   
   ////MSHIFTSBR
   	ELSIF (TMP_dSourceFile = 201) AND (TMP_dDestFile = 200) THEN
   		COP(N201[TMP_dSourceOffset], N200[TMP_dDestOffset], TMP_dNumValues);
   	ELSIF (TMP_dSourceFile = 202) AND (TMP_dDestFile = 200) THEN
   		COP(N202[TMP_dSourceOffset], N200[TMP_dDestOffset], TMP_dNumValues);
   	ELSIF (TMP_dSourceFile = 203) AND (TMP_dDestFile = 200) THEN
   		COP(N203[TMP_dSourceOffset], N200[TMP_dDestOffset], TMP_dNumValues);
   	ELSIF (TMP_dSourceFile = 204) AND (TMP_dDestFile = 200) THEN
   		COP(N204[TMP_dSourceOffset], N200[TMP_dDestOffset], TMP_dNumValues);
   	ELSIF (TMP_dSourceFile = 205) AND (TMP_dDestFile = 200) THEN
   		COP(N205[TMP_dSourceOffset], N200[TMP_dDestOffset], TMP_dNumValues);
   	ELSIF (TMP_dSourceFile = 206) AND (TMP_dDestFile = 200) THEN
   		COP(N206[TMP_dSourceOffset], N200[TMP_dDestOffset], TMP_dNumValues);
   	ELSIF (TMP_dSourceFile = 207) AND (TMP_dDestFile = 200) THEN
   		COP(N207[TMP_dSourceOffset], N200[TMP_dDestOffset], TMP_dNumValues);
   	ELSIF (TMP_dSourceFile = 208) AND (TMP_dDestFile = 200) THEN
   		COP(N208[TMP_dSourceOffset], N200[TMP_dDestOffset], TMP_dNumValues);
   	ELSIF (TMP_dSourceFile = 209) AND (TMP_dDestFile = 200) THEN
   		COP(N209[TMP_dSourceOffset], N200[TMP_dDestOffset], TMP_dNumValues);
   	ELSIF (TMP_dSourceFile = 210) AND (TMP_dDestFile = 200) THEN
   		COP(N210[TMP_dSourceOffset], N200[TMP_dDestOffset], TMP_dNumValues);
   	ELSIF (TMP_dSourceFile = 211) AND (TMP_dDestFile = 200) THEN
   		COP(N211[TMP_dSourceOffset], N200[TMP_dDestOffset], TMP_dNumValues);
   	ELSIF (TMP_dSourceFile = 212) AND (TMP_dDestFile = 200) THEN
   		COP(N212[TMP_dSourceOffset], N200[TMP_dDestOffset], TMP_dNumValues);
   	ELSIF (TMP_dSourceFile = 213) AND (TMP_dDestFile = 200) THEN
   		COP(N213[TMP_dSourceOffset], N200[TMP_dDestOffset], TMP_dNumValues);
   	ELSIF (TMP_dSourceFile = 214) AND (TMP_dDestFile = 200) THEN
   		COP(N214[TMP_dSourceOffset], N200[TMP_dDestOffset], TMP_dNumValues);
   	ELSIF (TMP_dSourceFile = 215) AND (TMP_dDestFile = 200) THEN
   		COP(N215[TMP_dSourceOffset], N200[TMP_dDestOffset], TMP_dNumValues);
   	ELSIF (TMP_dSourceFile = 216) AND (TMP_dDestFile = 200) THEN
   		COP(N216[TMP_dSourceOffset], N200[TMP_dDestOffset], TMP_dNumValues);
   	ELSIF (TMP_dSourceFile = 217) AND (TMP_dDestFile = 200) THEN
   		COP(N217[TMP_dSourceOffset], N200[TMP_dDestOffset], TMP_dNumValues);
   	ELSIF (TMP_dSourceFile = 218) AND (TMP_dDestFile = 200) THEN
   		COP(N218[TMP_dSourceOffset], N200[TMP_dDestOffset], TMP_dNumValues);
   
   	ELSIF (TMP_dSourceFile = 200) AND (TMP_dDestFile = 201) THEN
   		COP(N200[TMP_dSourceOffset], N201[TMP_dDestOffset], TMP_dNumValues);
   	ELSIF (TMP_dSourceFile = 200) AND (TMP_dDestFile = 202) THEN
   		COP(N200[TMP_dSourceOffset], N202[TMP_dDestOffset], TMP_dNumValues);
   	ELSIF (TMP_dSourceFile = 200) AND (TMP_dDestFile = 203) THEN
   		COP(N200[TMP_dSourceOffset], N203[TMP_dDestOffset], TMP_dNumValues);
   	ELSIF (TMP_dSourceFile = 200) AND (TMP_dDestFile = 204) THEN
   		COP(N200[TMP_dSourceOffset], N204[TMP_dDestOffset], TMP_dNumValues);
   	ELSIF (TMP_dSourceFile = 200) AND (TMP_dDestFile = 205) THEN
   		COP(N200[TMP_dSourceOffset], N205[TMP_dDestOffset], TMP_dNumValues);
   	ELSIF (TMP_dSourceFile = 200) AND (TMP_dDestFile = 206) THEN
   		COP(N200[TMP_dSourceOffset], N206[TMP_dDestOffset], TMP_dNumValues);
   	ELSIF (TMP_dSourceFile = 200) AND (TMP_dDestFile = 207) THEN
   		COP(N200[TMP_dSourceOffset], N207[TMP_dDestOffset], TMP_dNumValues);
   	ELSIF (TMP_dSourceFile = 200) AND (TMP_dDestFile = 208) THEN
   		COP(N200[TMP_dSourceOffset], N208[TMP_dDestOffset], TMP_dNumValues);
   	ELSIF (TMP_dSourceFile = 200) AND (TMP_dDestFile = 209) THEN
   		COP(N200[TMP_dSourceOffset], N209[TMP_dDestOffset], TMP_dNumValues);
   	ELSIF (TMP_dSourceFile = 200) AND (TMP_dDestFile = 210) THEN
   		COP(N200[TMP_dSourceOffset], N210[TMP_dDestOffset], TMP_dNumValues);
   	ELSIF (TMP_dSourceFile = 200) AND (TMP_dDestFile = 211) THEN
   		COP(N200[TMP_dSourceOffset], N211[TMP_dDestOffset], TMP_dNumValues);
   	ELSIF (TMP_dSourceFile = 200) AND (TMP_dDestFile = 212) THEN
   		COP(N200[TMP_dSourceOffset], N212[TMP_dDestOffset], TMP_dNumValues);
   	ELSIF (TMP_dSourceFile = 200) AND (TMP_dDestFile = 213) THEN
   		COP(N200[TMP_dSourceOffset], N213[TMP_dDestOffset], TMP_dNumValues);
   	ELSIF (TMP_dSourceFile = 200) AND (TMP_dDestFile = 214) THEN
   		COP(N200[TMP_dSourceOffset], N214[TMP_dDestOffset], TMP_dNumValues);
   	ELSIF (TMP_dSourceFile = 200) AND (TMP_dDestFile = 215) THEN
   		COP(N200[TMP_dSourceOffset], N215[TMP_dDestOffset], TMP_dNumValues);
   	ELSIF (TMP_dSourceFile = 200) AND (TMP_dDestFile = 216) THEN
   		COP(N200[TMP_dSourceOffset], N216[TMP_dDestOffset], TMP_dNumValues);
   	ELSIF (TMP_dSourceFile = 200) AND (TMP_dDestFile = 217) THEN
   		COP(N200[TMP_dSourceOffset], N217[TMP_dDestOffset], TMP_dNumValues);
   	ELSIF (TMP_dSourceFile = 200) AND (TMP_dDestFile = 218) THEN
   		COP(N200[TMP_dSourceOffset], N218[TMP_dDestOffset], TMP_dNumValues);
   
   
   ////////
   	ELSE
   		TMP_dErrSourceFile := TMP_dSourceFile;
   		TMP_dErrDestFile := TMP_dDestFile;
   	END_IF;
   *)
   
   RET(TMP_dErrSourceFile,TMP_dErrDestFile);
   
END_ROUTINE

ROUTINE _9_MCP_H   (* ladder *)
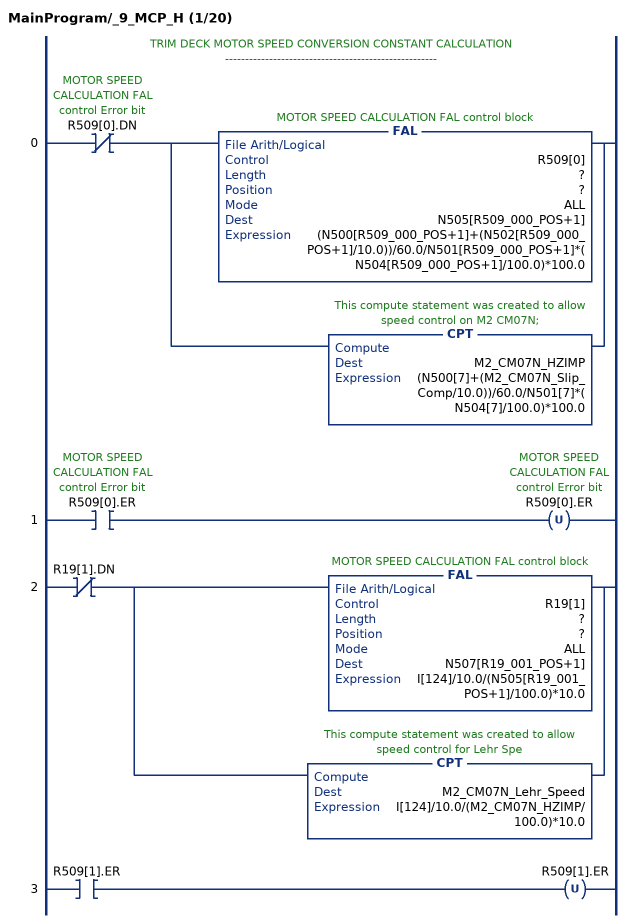
   // TRIM DECK MOTOR SPEED CONVERSION CONSTANT CALCULATION
   // -----------------------------------------------------
   0: XIO(R509[0].DN)[FAL(R509[0],?,?,ALL,N505[R509_000_POS+1],(N500[R509_000_POS+1]+(N502[R509_000_POS+1]/10.0))/60.0/N501[R509_000_POS+1]*(N504[R509_000_POS+1]/100.0)*100.0) ,CPT(M2_CM07N_HZIMP,(N500[7]+(M2_CM07N_Slip_Comp/10.0))/60.0/N501[7]*(N504[7]/100.0)*100.0) ];
   1: XIC(R509[0].ER)OTU(R509[0].ER);
   2: XIO(R19[1].DN)[FAL(R19[1],?,?,ALL,N507[R19_001_POS+1],I[124]/10.0/(N505[R19_001_POS+1]/100.0)*10.0) ,CPT(M2_CM07N_Lehr_Speed,I[124]/10.0/(M2_CM07N_HZIMP/100.0)*10.0) ];
   3: XIC(R509[1].ER)OTU(R509[1].ER);
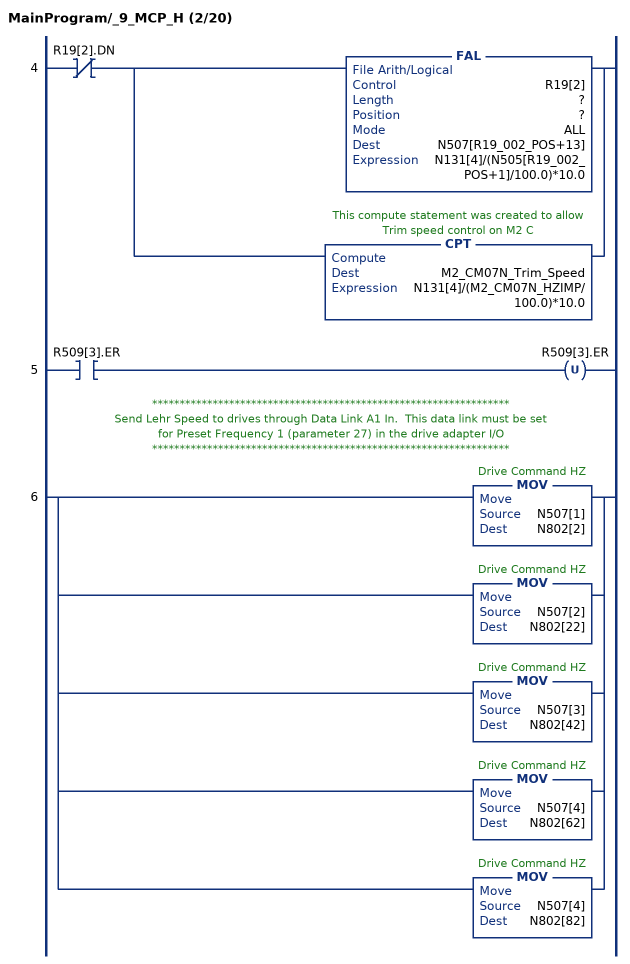
   4: XIO(R19[2].DN)[FAL(R19[2],?,?,ALL,N507[R19_002_POS+13],N131[4]/(N505[R19_002_POS+1]/100.0)*10.0) ,CPT(M2_CM07N_Trim_Speed,N131[4]/(M2_CM07N_HZIMP/100.0)*10.0) ];
   5: XIC(R509[3].ER)OTU(R509[3].ER);
   // *****************************************************************
   // Send Lehr Speed to drives through Data Link A1 In.  This data link must be set
   // for Preset Frequency 1 (parameter 27) in the drive adapter I/O
   // *****************************************************************
   6: [MOV(N507[1],N802[2]) ,MOV(N507[2],N802[22]) ,MOV(N507[3],N802[42]) ,MOV(N507[4],N802[62]) ,MOV(N507[4],N802[82]) ];
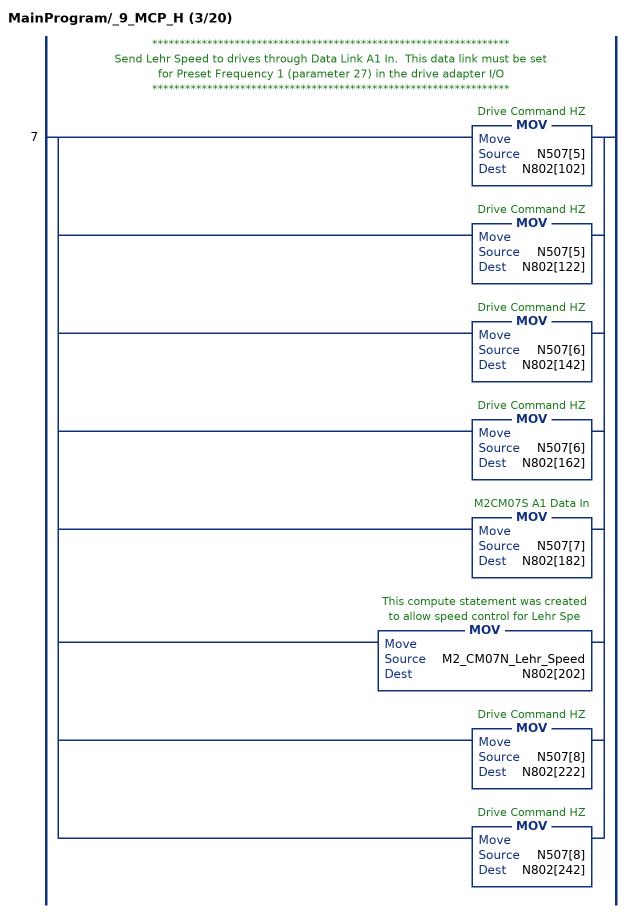
   // *****************************************************************
   // Send Lehr Speed to drives through Data Link A1 In.  This data link must be set
   // for Preset Frequency 1 (parameter 27) in the drive adapter I/O
   // *****************************************************************
   7: [MOV(N507[5],N802[102]) ,MOV(N507[5],N802[122]) ,MOV(N507[6],N802[142]) ,MOV(N507[6],N802[162]) ,MOV(N507[7],N802[182]) ,MOV(M2_CM07N_Lehr_Speed,N802[202]) ,MOV(N507[8],N802[222]) ,MOV(N507[8],N802[242]) ];
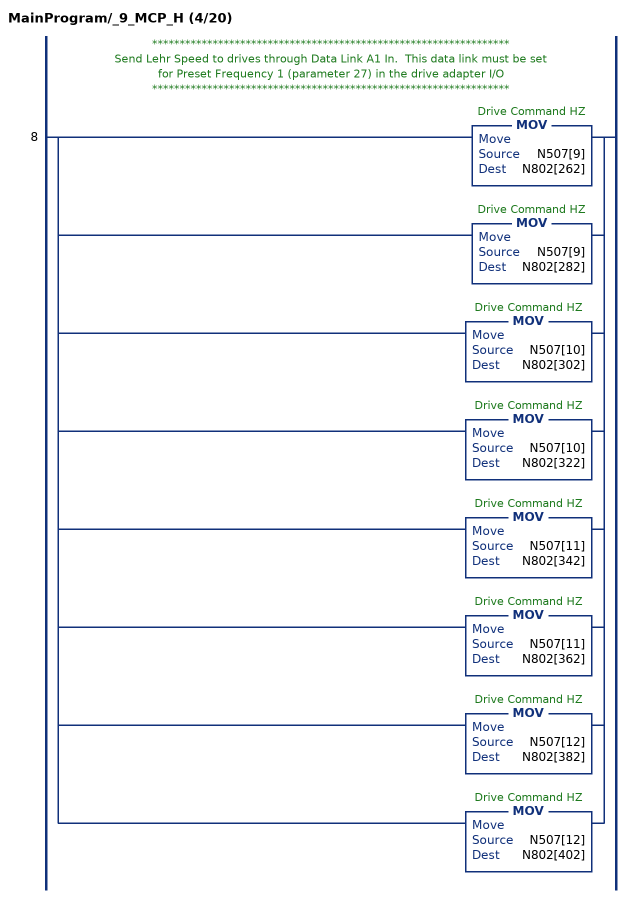
   // *****************************************************************
   // Send Lehr Speed to drives through Data Link A1 In.  This data link must be set
   // for Preset Frequency 1 (parameter 27) in the drive adapter I/O
   // *****************************************************************
   8: [MOV(N507[9],N802[262]) ,MOV(N507[9],N802[282]) ,MOV(N507[10],N802[302]) ,MOV(N507[10],N802[322]) ,MOV(N507[11],N802[342]) ,MOV(N507[11],N802[362]) ,MOV(N507[12],N802[382]) ,MOV(N507[12],N802[402]) ];
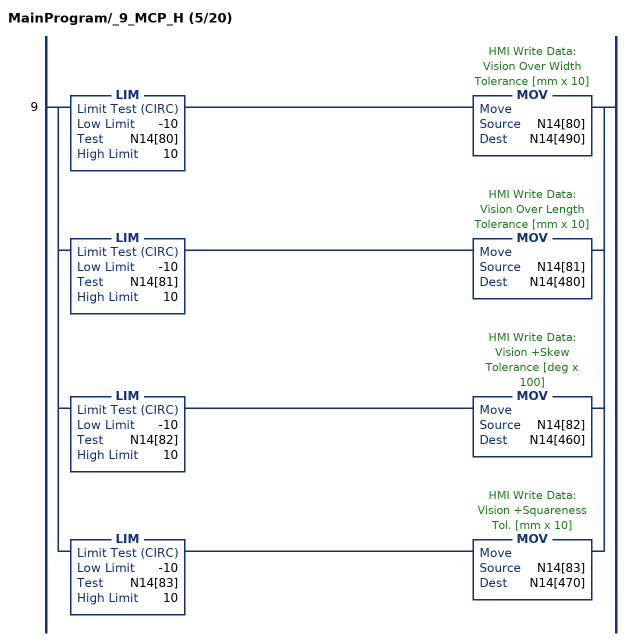
   9: [LIM(-10,N14[80],10) MOV(N14[80],N14[490]) ,LIM(-10,N14[81],10) MOV(N14[81],N14[480]) ,LIM(-10,N14[82],10) MOV(N14[82],N14[460]) ,LIM(-10,N14[83],10) MOV(N14[83],N14[470]) ];
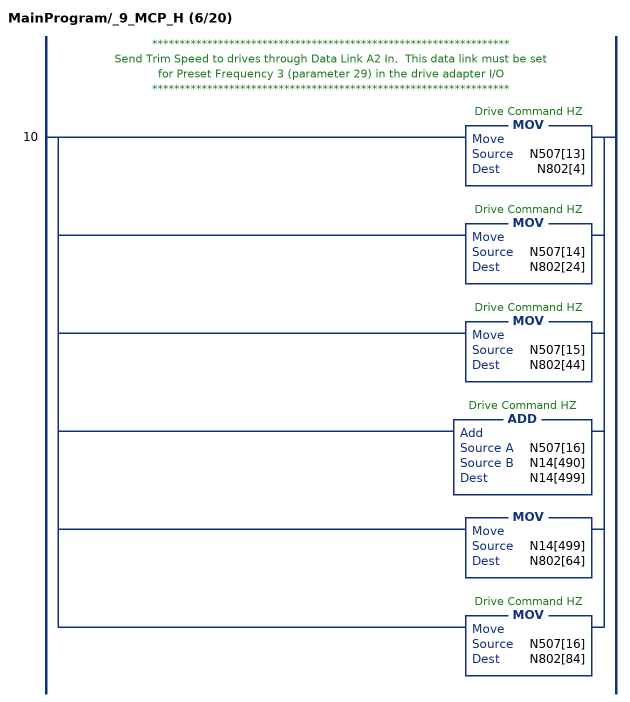
   // *****************************************************************
   // Send Trim Speed to drives through Data Link A2 In.  This data link must be set
   // for Preset Frequency 3 (parameter 29) in the drive adapter I/O
   // *****************************************************************
   10: [MOV(N507[13],N802[4]) ,MOV(N507[14],N802[24]) ,MOV(N507[15],N802[44]) ,ADD(N507[16],N14[490],N14[499]) ,MOV(N14[499],N802[64]) ,MOV(N507[16],N802[84]) ];
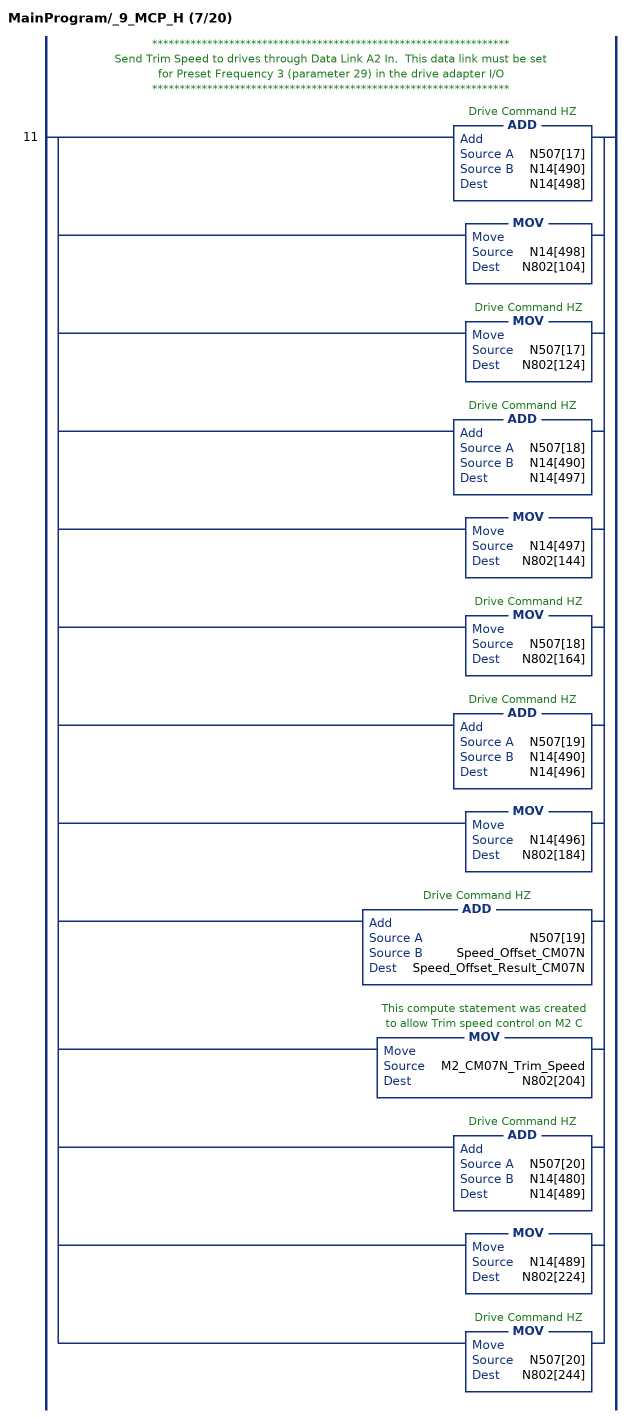
   // *****************************************************************
   // Send Trim Speed to drives through Data Link A2 In.  This data link must be set
   // for Preset Frequency 3 (parameter 29) in the drive adapter I/O
   // *****************************************************************
   11: [ADD(N507[17],N14[490],N14[498]) ,MOV(N14[498],N802[104]) ,MOV(N507[17],N802[124]) ,ADD(N507[18],N14[490],N14[497]) ,MOV(N14[497],N802[144]) ,MOV(N507[18],N802[164]) ,ADD(N507[19],N14[490],N14[496]) ,MOV(N14[496],N802[184]) ,ADD(N507[19],Speed_Offset_CM07N,Speed_Offset_Result_CM07N) ,MOV(M2_CM07N_Trim_Speed,N802[204]) ,ADD(N507[20],N14[480],N14[489]) ,MOV(N14[489],N802[224]) ,MOV(N507[20],N802[244]) ];
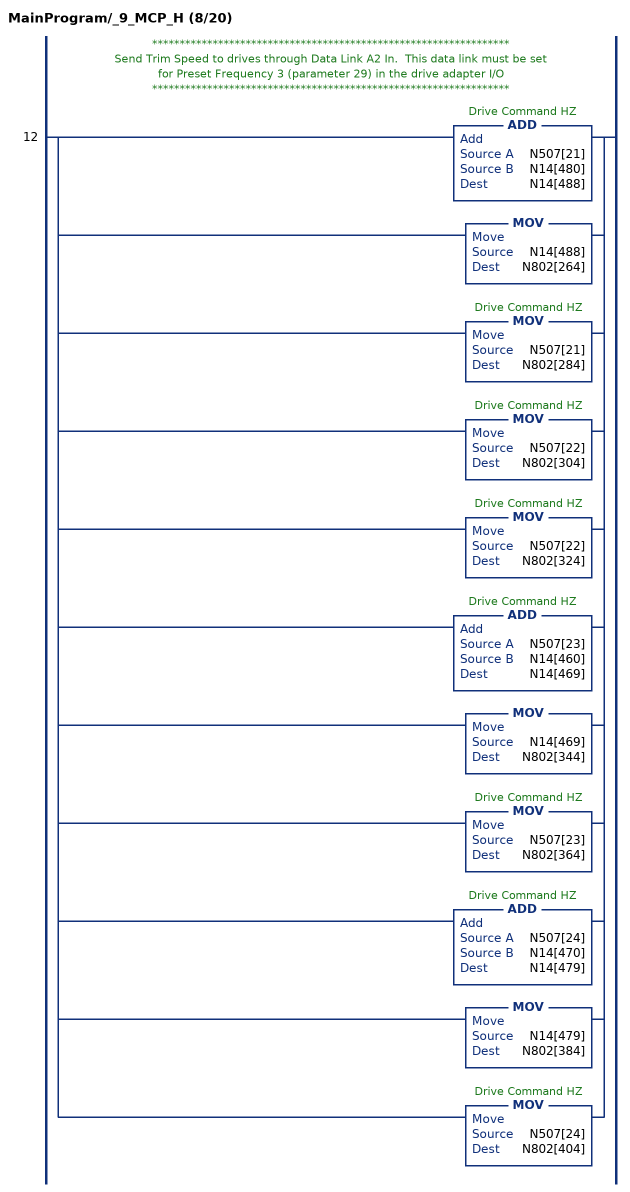
   // *****************************************************************
   // Send Trim Speed to drives through Data Link A2 In.  This data link must be set
   // for Preset Frequency 3 (parameter 29) in the drive adapter I/O
   // *****************************************************************
   12: [ADD(N507[21],N14[480],N14[488]) ,MOV(N14[488],N802[264]) ,MOV(N507[21],N802[284]) ,MOV(N507[22],N802[304]) ,MOV(N507[22],N802[324]) ,ADD(N507[23],N14[460],N14[469]) ,MOV(N14[469],N802[344]) ,MOV(N507[23],N802[364]) ,ADD(N507[24],N14[470],N14[479]) ,MOV(N14[479],N802[384]) ,MOV(N507[24],N802[404]) ];
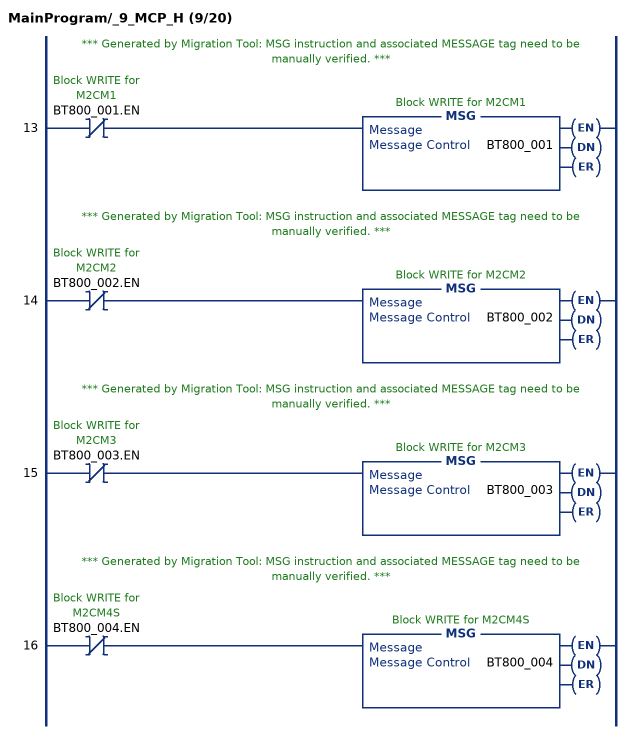
   // *** Generated by Migration Tool: MSG instruction and associated MESSAGE tag need to be manually verified. ***
   13: XIO(BT800_001.EN)MSG(BT800_001);
   // *** Generated by Migration Tool: MSG instruction and associated MESSAGE tag need to be manually verified. ***
   14: XIO(BT800_002.EN)MSG(BT800_002);
   // *** Generated by Migration Tool: MSG instruction and associated MESSAGE tag need to be manually verified. ***
   15: XIO(BT800_003.EN)MSG(BT800_003);
   // *** Generated by Migration Tool: MSG instruction and associated MESSAGE tag need to be manually verified. ***
   16: XIO(BT800_004.EN)MSG(BT800_004);
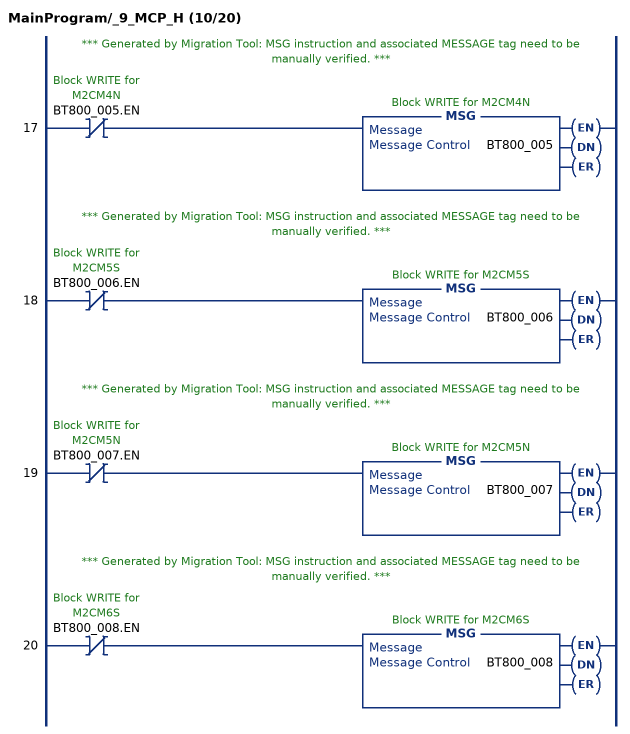
   // *** Generated by Migration Tool: MSG instruction and associated MESSAGE tag need to be manually verified. ***
   17: XIO(BT800_005.EN)MSG(BT800_005);
   // *** Generated by Migration Tool: MSG instruction and associated MESSAGE tag need to be manually verified. ***
   18: XIO(BT800_006.EN)MSG(BT800_006);
   // *** Generated by Migration Tool: MSG instruction and associated MESSAGE tag need to be manually verified. ***
   19: XIO(BT800_007.EN)MSG(BT800_007);
   // *** Generated by Migration Tool: MSG instruction and associated MESSAGE tag need to be manually verified. ***
   20: XIO(BT800_008.EN)MSG(BT800_008);
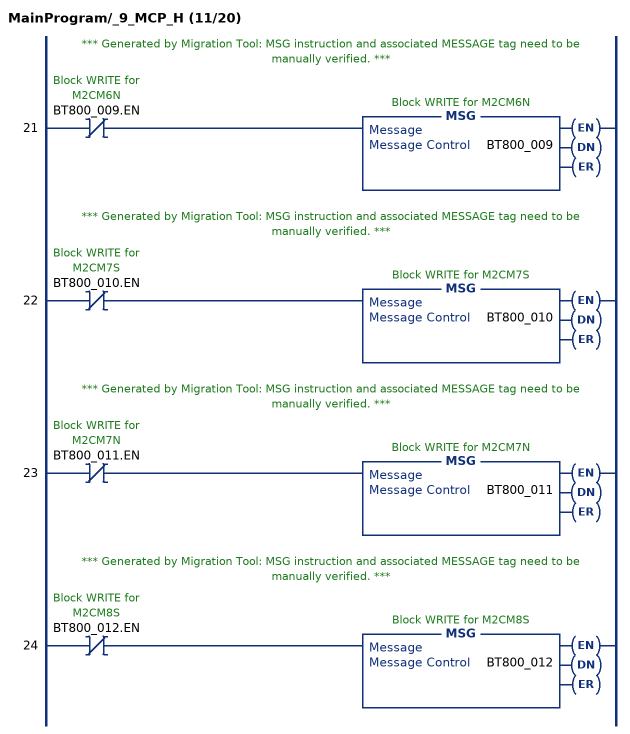
   // *** Generated by Migration Tool: MSG instruction and associated MESSAGE tag need to be manually verified. ***
   21: XIO(BT800_009.EN)MSG(BT800_009);
   // *** Generated by Migration Tool: MSG instruction and associated MESSAGE tag need to be manually verified. ***
   22: XIO(BT800_010.EN)MSG(BT800_010);
   // *** Generated by Migration Tool: MSG instruction and associated MESSAGE tag need to be manually verified. ***
   23: XIO(BT800_011.EN)MSG(BT800_011);
   // *** Generated by Migration Tool: MSG instruction and associated MESSAGE tag need to be manually verified. ***
   24: XIO(BT800_012.EN)MSG(BT800_012);
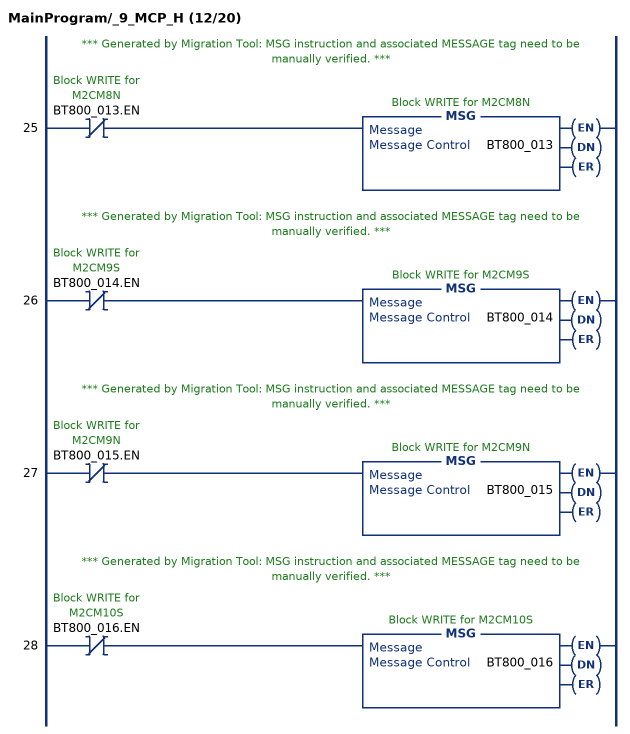
   // *** Generated by Migration Tool: MSG instruction and associated MESSAGE tag need to be manually verified. ***
   25: XIO(BT800_013.EN)MSG(BT800_013);
   // *** Generated by Migration Tool: MSG instruction and associated MESSAGE tag need to be manually verified. ***
   26: XIO(BT800_014.EN)MSG(BT800_014);
   // *** Generated by Migration Tool: MSG instruction and associated MESSAGE tag need to be manually verified. ***
   27: XIO(BT800_015.EN)MSG(BT800_015);
   // *** Generated by Migration Tool: MSG instruction and associated MESSAGE tag need to be manually verified. ***
   28: XIO(BT800_016.EN)MSG(BT800_016);
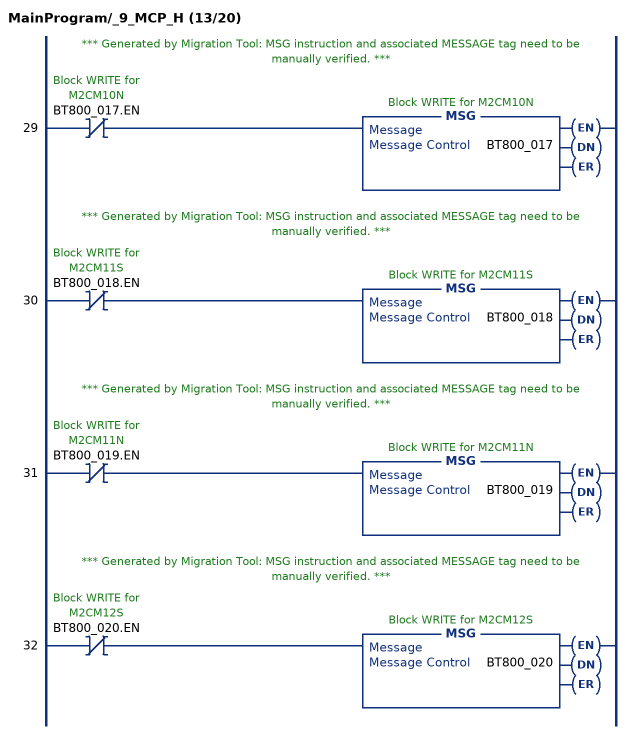
   // *** Generated by Migration Tool: MSG instruction and associated MESSAGE tag need to be manually verified. ***
   29: XIO(BT800_017.EN)MSG(BT800_017);
   // *** Generated by Migration Tool: MSG instruction and associated MESSAGE tag need to be manually verified. ***
   30: XIO(BT800_018.EN)MSG(BT800_018);
   // *** Generated by Migration Tool: MSG instruction and associated MESSAGE tag need to be manually verified. ***
   31: XIO(BT800_019.EN)MSG(BT800_019);
   // *** Generated by Migration Tool: MSG instruction and associated MESSAGE tag need to be manually verified. ***
   32: XIO(BT800_020.EN)MSG(BT800_020);
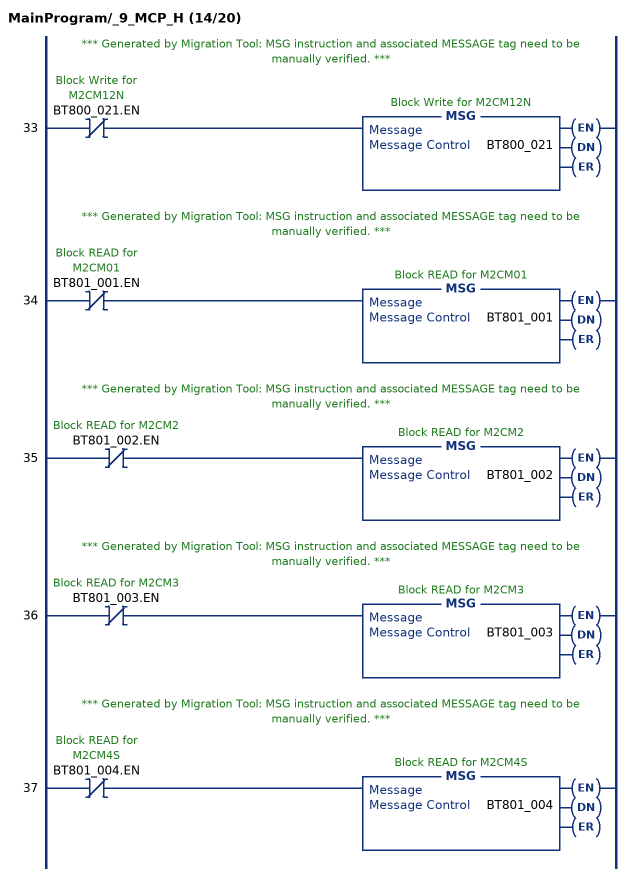
   // *** Generated by Migration Tool: MSG instruction and associated MESSAGE tag need to be manually verified. ***
   33: XIO(BT800_021.EN)MSG(BT800_021);
   // *** Generated by Migration Tool: MSG instruction and associated MESSAGE tag need to be manually verified. ***
   34: XIO(BT801_001.EN)MSG(BT801_001);
   // *** Generated by Migration Tool: MSG instruction and associated MESSAGE tag need to be manually verified. ***
   35: XIO(BT801_002.EN)MSG(BT801_002);
   // *** Generated by Migration Tool: MSG instruction and associated MESSAGE tag need to be manually verified. ***
   36: XIO(BT801_003.EN)MSG(BT801_003);
   // *** Generated by Migration Tool: MSG instruction and associated MESSAGE tag need to be manually verified. ***
   37: XIO(BT801_004.EN)MSG(BT801_004);
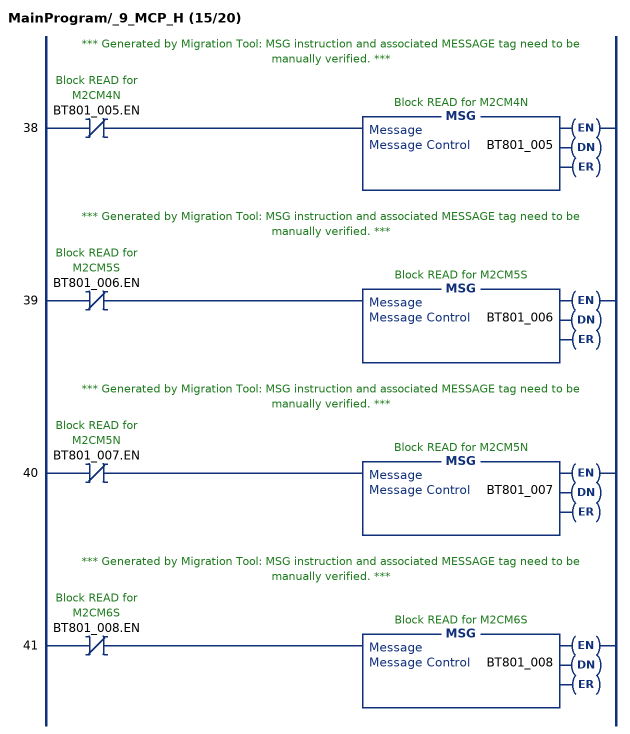
   // *** Generated by Migration Tool: MSG instruction and associated MESSAGE tag need to be manually verified. ***
   38: XIO(BT801_005.EN)MSG(BT801_005);
   // *** Generated by Migration Tool: MSG instruction and associated MESSAGE tag need to be manually verified. ***
   39: XIO(BT801_006.EN)MSG(BT801_006);
   // *** Generated by Migration Tool: MSG instruction and associated MESSAGE tag need to be manually verified. ***
   40: XIO(BT801_007.EN)MSG(BT801_007);
   // *** Generated by Migration Tool: MSG instruction and associated MESSAGE tag need to be manually verified. ***
   41: XIO(BT801_008.EN)MSG(BT801_008);
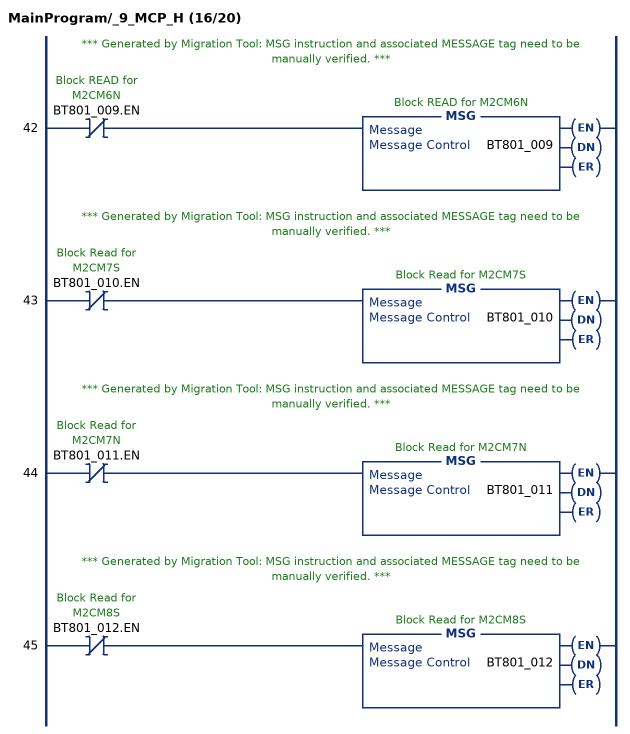
   // *** Generated by Migration Tool: MSG instruction and associated MESSAGE tag need to be manually verified. ***
   42: XIO(BT801_009.EN)MSG(BT801_009);
   // *** Generated by Migration Tool: MSG instruction and associated MESSAGE tag need to be manually verified. ***
   43: XIO(BT801_010.EN)MSG(BT801_010);
   // *** Generated by Migration Tool: MSG instruction and associated MESSAGE tag need to be manually verified. ***
   44: XIO(BT801_011.EN)MSG(BT801_011);
   // *** Generated by Migration Tool: MSG instruction and associated MESSAGE tag need to be manually verified. ***
   45: XIO(BT801_012.EN)MSG(BT801_012);
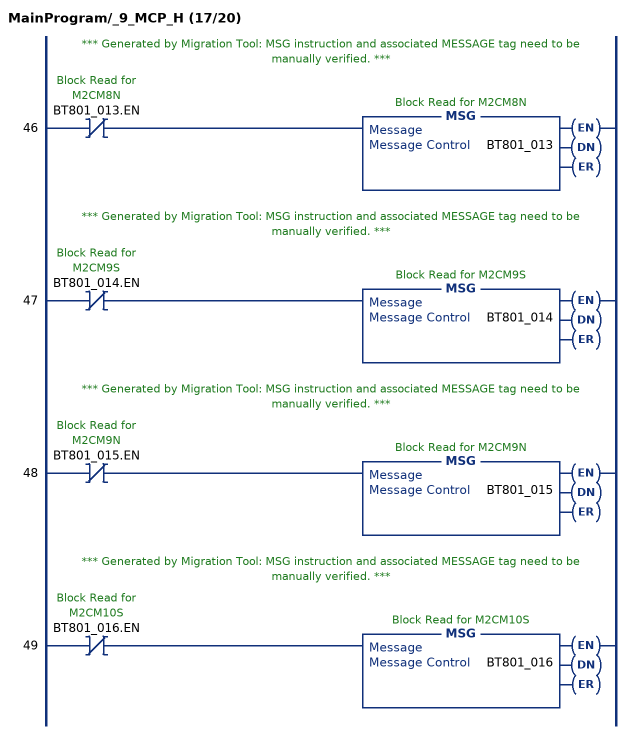
   // *** Generated by Migration Tool: MSG instruction and associated MESSAGE tag need to be manually verified. ***
   46: XIO(BT801_013.EN)MSG(BT801_013);
   // *** Generated by Migration Tool: MSG instruction and associated MESSAGE tag need to be manually verified. ***
   47: XIO(BT801_014.EN)MSG(BT801_014);
   // *** Generated by Migration Tool: MSG instruction and associated MESSAGE tag need to be manually verified. ***
   48: XIO(BT801_015.EN)MSG(BT801_015);
   // *** Generated by Migration Tool: MSG instruction and associated MESSAGE tag need to be manually verified. ***
   49: XIO(BT801_016.EN)MSG(BT801_016);
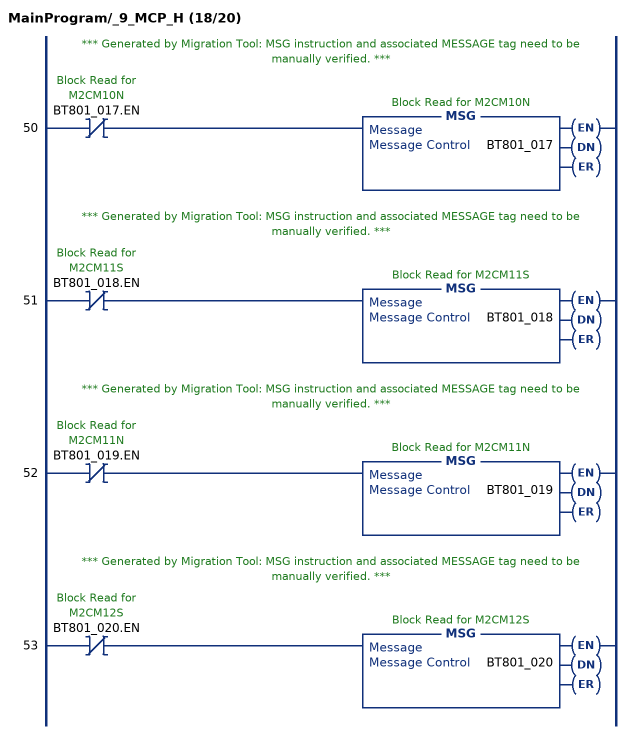
   // *** Generated by Migration Tool: MSG instruction and associated MESSAGE tag need to be manually verified. ***
   50: XIO(BT801_017.EN)MSG(BT801_017);
   // *** Generated by Migration Tool: MSG instruction and associated MESSAGE tag need to be manually verified. ***
   51: XIO(BT801_018.EN)MSG(BT801_018);
   // *** Generated by Migration Tool: MSG instruction and associated MESSAGE tag need to be manually verified. ***
   52: XIO(BT801_019.EN)MSG(BT801_019);
   // *** Generated by Migration Tool: MSG instruction and associated MESSAGE tag need to be manually verified. ***
   53: XIO(BT801_020.EN)MSG(BT801_020);
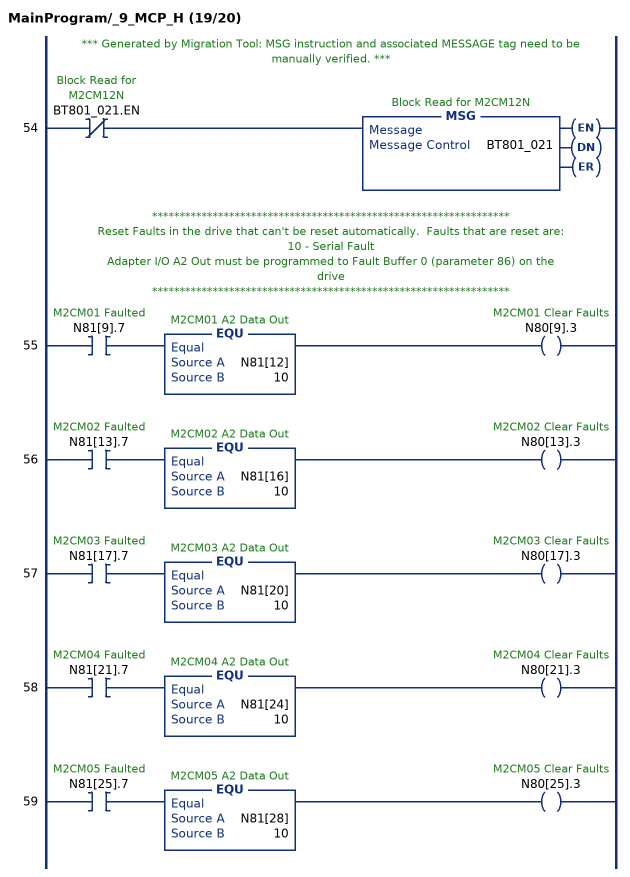
   // *** Generated by Migration Tool: MSG instruction and associated MESSAGE tag need to be manually verified. ***
   54: XIO(BT801_021.EN)MSG(BT801_021);
   // *****************************************************************
   // Reset Faults in the drive that can't be reset automatically.  Faults that are reset are:
   //  10 - Serial Fault
   // Adapter I/O A2 Out must be programmed to Fault Buffer 0 (parameter 86) on the
   // drive
   // *****************************************************************
   55: XIC(N81[9].7)EQU(N81[12],10)OTE(N80[9].3);
   56: XIC(N81[13].7)EQU(N81[16],10)OTE(N80[13].3);
   57: XIC(N81[17].7)EQU(N81[20],10)OTE(N80[17].3);
   58: XIC(N81[21].7)EQU(N81[24],10)OTE(N80[21].3);
   59: XIC(N81[25].7)EQU(N81[28],10)OTE(N80[25].3);
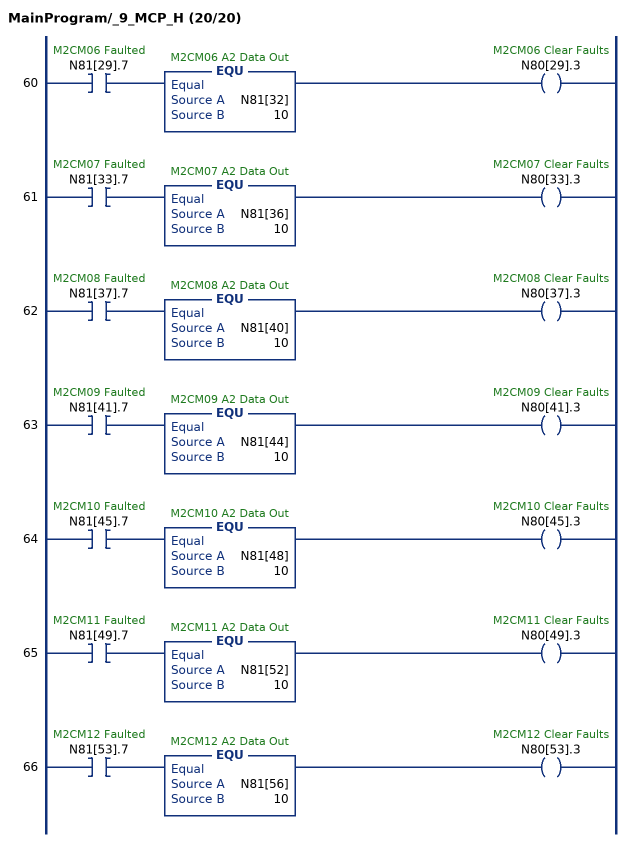
   60: XIC(N81[29].7)EQU(N81[32],10)OTE(N80[29].3);
   61: XIC(N81[33].7)EQU(N81[36],10)OTE(N80[33].3);
   62: XIC(N81[37].7)EQU(N81[40],10)OTE(N80[37].3);
   63: XIC(N81[41].7)EQU(N81[44],10)OTE(N80[41].3);
   64: XIC(N81[45].7)EQU(N81[48],10)OTE(N80[45].3);
   65: XIC(N81[49].7)EQU(N81[52],10)OTE(N80[49].3);
   66: XIC(N81[53].7)EQU(N81[56],10)OTE(N80[53].3);
END_ROUTINE
